VERSION : 0.1
   VAR_INPUT
      IN_xCycleON : Bool;   // Cycle ON
      IN_xCycleONDel : Bool;   // Delayed cycle ON signal
      IN_xResetAlarms : Bool;   // Reset alarms
      IN_xFaultsEnabled : Bool;   // Faults enabled
      IN_xAccelation : Bool;
      IN_rgtMotorConfig : "UDT_MotorConfig";
   END_VAR
   VAR
      ST_xCondOkMan : Bool;   // Manual condition Ok
      ST_xManualMode : Bool;   // Manual mode
      ST_xMachineAnomaly : Bool;   // Machine anomaly
      ST_xStoppingFaults : Bool;   // Stopping fault
      ST_xFaults : Bool;   // Fault
      ST_xWarnings : Bool;   // Warnings
      ST_xConditionOkStopCycle : Bool;   // Condition ok stop cycle
      ST_xOutputEnable : Bool;   // Output enable
      ST_xFeedbackRotation : Bool;   // Feedback rotation
      ST_xPowerUnitSwitchOnRequest : Bool;   // Power unit switch on request
      INPUT_xLocalSwitch : Bool;   // Input local safety switch
      INPUT_xQFMotorFan : Bool;   // Input motor fan protection
      INPUT_xMotorThermalProbe : Bool;   // Input motor thermal probe
      INPUT_xPowerModuleOn : Bool;   // Input power module switched on
      INPUT_dMagnitude : Int;   // Input magnitude value from drive
      INPUT_dTorque : Int;   // Input torque value from drive
      AUX_dReqSpeed_mm_min : DInt := 0;   // Conveyor requested speed [mm/min]
      AUX_dlimitTorqueCorrection : DInt := 0;   // Limit Torque [mm/min]
      tmON_DelayReadyToMove : "UDT_IECTON_V1.00";   // Delay ready to move
      tmON_FeedbackTimeOut : "UDT_IECTON_V1.00";   // Feedback Time out
      tmOF_DriveEnable : "UDT_IECTON_V1.00";   // Drive enable dealy
      AUX_rgtSinamicsIDB : "SINAMICS_LinearPos_ControlTorque";
      tHMR : Struct   // {[Unit]|[Scada Unit]|[LowLimit]|[HigLimit]|[Acces]}
         xManualCommandEnabled : Bool;   // Manual Command enabled {x|x|x|x|O}
         dState : DInt;   // State Conveyor (1=No anomaly, 3=Run, 7=Anomaly) {x|x|x|x|O}
         dMagnitudeCurrent : DInt;   // Magnitude Current [mA] {mA|A|x|x|O}
         dTorque : DInt;   // Torque value [mN] {mN|N|x|x|O}
         dSpeedFeedback : DInt;   // Speed Feedback [mm/min] {mm/min|m/min|x|x|O}
         tManCmd : Struct
            xFdbkRunFw : Bool;   // Motor Rotation Enabled FW {x|x|x|x|O}
         END_STRUCT;
      END_STRUCT;
      tHMW : Struct   // {[Unit]|[Scada Unit]|[LowLimit]|[HigLimit]|[Acces]}
         xEnableManualCommand : Bool;   // Enable Manual command {x|x|x|x|O}
         dSpeedCorrection : DInt;   // Speed Correction[‰] {‰|%|-2|2|M}
         dCurrentLimit : DInt;   // Current limit [‰] {‰|%|0|200|M}
         tManCmd : Struct
            xRunFw : Bool;   // Rotation FW {x|x|x|x|O}
         END_STRUCT;
      END_STRUCT;
      tALM : Struct   // HMI Alarms
         tS : Struct   // Stopping faults
            xLocalSafetySwitch : Bool;   // Local Safety Switch
            xFeedbackError : Bool;   // Feedback Error
            xDriveError : Bool;   // Drive Error
            xMotorFanProtection : Bool;   // Motor Fan protection
            xMotorThermalProbe : Bool;   // Motor Thermal Probe
            xSpare_5 : Bool;
            xSpare_6 : Bool;
            xSpare_7 : Bool;
            xSpare_8 : Bool;
            xSpare_9 : Bool;
            xSpare_10 : Bool;
            xSpare_11 : Bool;
            xSpare_12 : Bool;
            xSpare_13 : Bool;
            xSpare_14 : Bool;
            xSpare_15 : Bool;
            xSpare_16 : Bool;
            xSpare_17 : Bool;
            xSpare_18 : Bool;
            xSpare_19 : Bool;
            xSpare_20 : Bool;
            xSpare_21 : Bool;
            xSpare_22 : Bool;
            xSpare_23 : Bool;
            xSpare_24 : Bool;
            xSpare_25 : Bool;
            xSpare_26 : Bool;
            xSpare_27 : Bool;
            xSpare_28 : Bool;
            xSpare_29 : Bool;
            xSpare_30 : Bool;
            xSpare_31 : Bool;
         END_STRUCT;
         tF : Struct   // Faults
            xSpare_0 : Bool;
            xSpare_1 : Bool;
            xSpare_2 : Bool;
            xSpare_3 : Bool;
            xSpare_4 : Bool;
            xSpare_5 : Bool;
            xSpare_6 : Bool;
            xSpare_7 : Bool;
            xSpare_8 : Bool;
            xSpare_9 : Bool;
            xSpare_10 : Bool;
            xSpare_11 : Bool;
            xSpare_12 : Bool;
            xSpare_13 : Bool;
            xSpare_14 : Bool;
            xSpare_15 : Bool;
            xSpare_16 : Bool;
            xSpare_17 : Bool;
            xSpare_18 : Bool;
            xSpare_19 : Bool;
            xSpare_20 : Bool;
            xSpare_21 : Bool;
            xSpare_22 : Bool;
            xSpare_23 : Bool;
            xSpare_24 : Bool;
            xSpare_25 : Bool;
            xSpare_26 : Bool;
            xSpare_27 : Bool;
            xSpare_28 : Bool;
            xSpare_29 : Bool;
            xSpare_30 : Bool;
            xSpare_31 : Bool;
         END_STRUCT;
         tW : Struct   // Warnings
            xSpare_0 : Bool;
            xSpare_1 : Bool;
            xSpare_2 : Bool;
            xSpare_3 : Bool;
            xSpare_4 : Bool;
            xSpare_5 : Bool;
            xSpare_6 : Bool;
            xSpare_7 : Bool;
            xSpare_8 : Bool;
            xSpare_9 : Bool;
            xSpare_10 : Bool;
            xSpare_11 : Bool;
            xSpare_12 : Bool;
            xSpare_13 : Bool;
            xSpare_14 : Bool;
            xSpare_15 : Bool;
            xSpare_16 : Bool;
            xSpare_17 : Bool;
            xSpare_18 : Bool;
            xSpare_19 : Bool;
            xSpare_20 : Bool;
            xSpare_21 : Bool;
            xSpare_22 : Bool;
            xSpare_23 : Bool;
            xSpare_24 : Bool;
            xSpare_25 : Bool;
            xSpare_26 : Bool;
            xSpare_27 : Bool;
            xSpare_28 : Bool;
            xSpare_29 : Bool;
            xSpare_30 : Bool;
            xSpare_31 : Bool;
         END_STRUCT;
      END_STRUCT;
   END_VAR
   VAR_TEMP
      TMP_dIndex : DInt;
      TMP_dwValue : DWord;
      TMP_iRetVal : Int;
      TMP_xDriveRun : Bool;
      TMP_xDriveEnable : Bool;
   END_VAR
   VAR_TEMP   // added for the SCL form of the ladder/FBD networks
      _w1 : Bool;
   END_VAR
BEGIN

REGION Network 1: #####_MATCH_#####
END_REGION

REGION Network 2: Feedback roller rotation
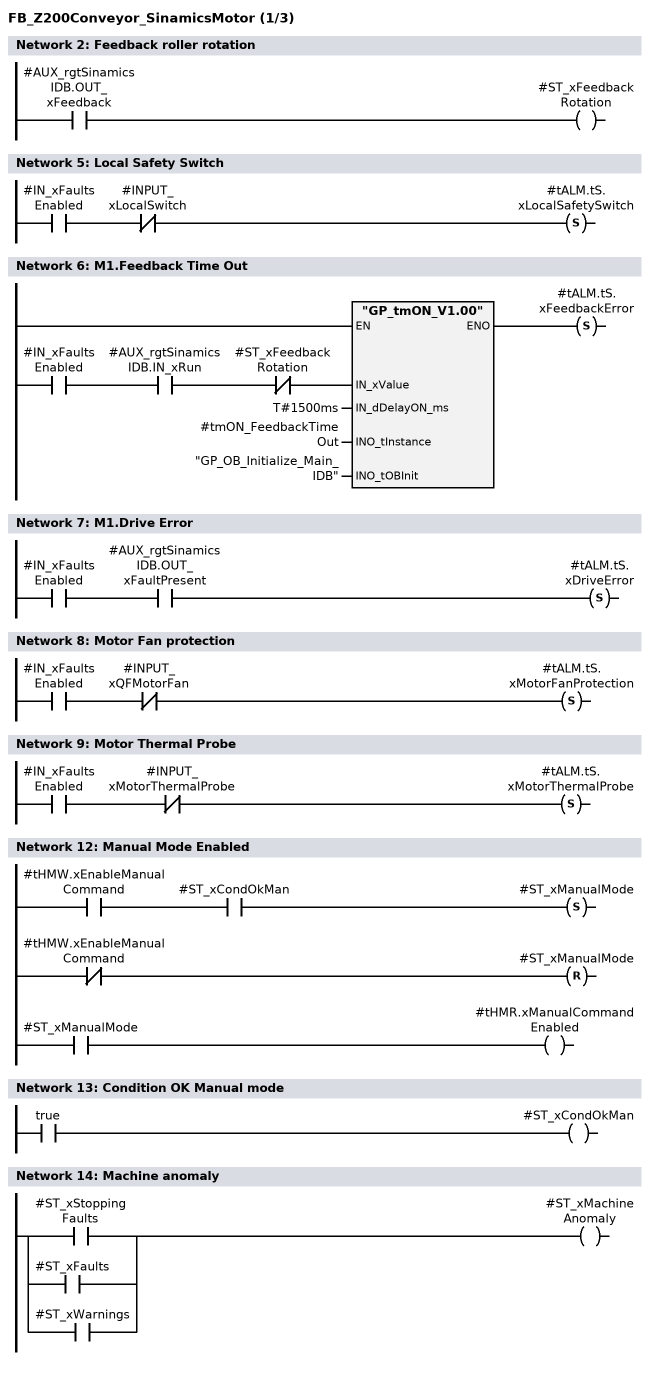
   RUNG wire#powerrail
      Contact( #AUX_rgtSinamicsIDB.OUT_xFeedback )
      Coil( #ST_xFeedbackRotation )
   END_RUNG
   // the same network as SCL:
   #ST_xFeedbackRotation := #AUX_rgtSinamicsIDB.OUT_xFeedback;
END_REGION

REGION Network 3: ####_ALARMS_####
END_REGION

REGION Network 4 (SCL): Reset alarms
   IF #IN_xResetAlarms THEN

       #TMP_dwValue := 0;

       SCATTER(IN:=#TMP_dwValue,
               OUT=>#tALM.tS);

       SCATTER(IN:=#TMP_dwValue,
               OUT=>#tALM.tF);

       SCATTER(IN:=#TMP_dwValue,
               OUT=>#tALM.tW);


   END_IF;
END_REGION

REGION Network 5: Local Safety Switch
   RUNG wire#powerrail
      Contact( #IN_xFaultsEnabled )
      I_Contact( #INPUT_xLocalSwitch )
      S_Coil( #tALM.tS.xLocalSafetySwitch )
   END_RUNG
   // the same network as SCL:
   IF #IN_xFaultsEnabled AND NOT #INPUT_xLocalSwitch THEN #tALM.tS.xLocalSafetySwitch := TRUE; END_IF;
END_REGION

REGION Network 6: M1.Feedback Time Out
   RUNG wire#powerrail
      "GP_tmON_V1.00"(IN_xValue := wire#w1, IN_dDelayON_ms := T#1500ms, INO_tInstance := #tmON_FeedbackTimeOut, INO_tOBInit := "GP_OB_Initialize_Main_IDB")
      S_Coil( #tALM.tS.xFeedbackError )
   END_RUNG
   RUNG wire#powerrail
      Contact( #IN_xFaultsEnabled )
      Contact( #AUX_rgtSinamicsIDB.IN_xRun )
      I_Contact( #ST_xFeedbackRotation )
   END_RUNG wire#w1
   // the same network as SCL:
   "GP_tmON_V1.00"(IN_xValue := #IN_xFaultsEnabled AND #AUX_rgtSinamicsIDB.IN_xRun AND NOT #ST_xFeedbackRotation,
                   IN_dDelayON_ms := T#1500ms,
                   INO_tInstance := #tmON_FeedbackTimeOut,
                   INO_tOBInit := "GP_OB_Initialize_Main_IDB",
                   ENO => #_w1);
   IF #_w1 THEN #tALM.tS.xFeedbackError := TRUE; END_IF;
END_REGION

REGION Network 7: M1.Drive Error
   RUNG wire#powerrail
      Contact( #IN_xFaultsEnabled )
      Contact( #AUX_rgtSinamicsIDB.OUT_xFaultPresent )
      S_Coil( #tALM.tS.xDriveError )
   END_RUNG
   // the same network as SCL:
   IF #IN_xFaultsEnabled AND #AUX_rgtSinamicsIDB.OUT_xFaultPresent THEN #tALM.tS.xDriveError := TRUE; END_IF;
END_REGION

REGION Network 8: Motor Fan protection
   RUNG wire#powerrail
      Contact( #IN_xFaultsEnabled )
      I_Contact( #INPUT_xQFMotorFan )
      S_Coil( #tALM.tS.xMotorFanProtection )
   END_RUNG
   // the same network as SCL:
   IF #IN_xFaultsEnabled AND NOT #INPUT_xQFMotorFan THEN #tALM.tS.xMotorFanProtection := TRUE; END_IF;
END_REGION

REGION Network 9: Motor Thermal Probe
   RUNG wire#powerrail
      Contact( #IN_xFaultsEnabled )
      I_Contact( #INPUT_xMotorThermalProbe )
      S_Coil( #tALM.tS.xMotorThermalProbe )
   END_RUNG
   // the same network as SCL:
   IF #IN_xFaultsEnabled AND NOT #INPUT_xMotorThermalProbe THEN #tALM.tS.xMotorThermalProbe := TRUE; END_IF;
END_REGION

REGION Network 10 (SCL): Calculate general statuses
   GATHER(IN:=#tALM.tS,
          OUT=>#TMP_dwValue);

   IF #TMP_dwValue <> 0 THEN
       #ST_xStoppingFaults := TRUE;
   ELSE
       #ST_xStoppingFaults := FALSE;
   END_IF;

   GATHER(IN:=#tALM.tF,
          OUT=>#TMP_dwValue);

   IF #TMP_dwValue <> 0 THEN
       #ST_xFaults := TRUE;
   ELSE
       #ST_xFaults := FALSE;
   END_IF;

   GATHER(IN:=#tALM.tW,
          OUT=>#TMP_dwValue);

   IF #TMP_dwValue <> 0 THEN
       #ST_xWarnings := TRUE;
   ELSE
       #ST_xWarnings := FALSE;
   END_IF;
END_REGION

REGION Network 11: #####_HMI_LOGICS_#####
END_REGION

REGION Network 12: Manual Mode Enabled
   RUNG wire#powerrail
      Contact( #tHMW.xEnableManualCommand )
      Contact( #ST_xCondOkMan )
      S_Coil( #ST_xManualMode )
   END_RUNG
   RUNG wire#powerrail
      I_Contact( #tHMW.xEnableManualCommand )
      R_Coil( #ST_xManualMode )
   END_RUNG
   RUNG wire#powerrail
      Contact( #ST_xManualMode )
      Coil( #tHMR.xManualCommandEnabled )
   END_RUNG
   // the same network as SCL:
   IF #tHMW.xEnableManualCommand AND #ST_xCondOkMan THEN #ST_xManualMode := TRUE; END_IF;
   IF NOT #tHMW.xEnableManualCommand THEN #ST_xManualMode := FALSE; END_IF;
   #tHMR.xManualCommandEnabled := #ST_xManualMode;
END_REGION

REGION Network 13: Condition OK Manual mode
   RUNG wire#powerrail
      Contact( true )
      Coil( #ST_xCondOkMan )
   END_RUNG
   // the same network as SCL:
   #ST_xCondOkMan := true;
END_REGION

REGION Network 14: Machine anomaly
   RUNG wire#powerrail
      Contact( #ST_xStoppingFaults )
      wire#w1
      Coil( #ST_xMachineAnomaly )
   END_RUNG
   RUNG wire#powerrail
      Contact( #ST_xFaults )
   END_RUNG wire#w1
   RUNG wire#powerrail
      Contact( #ST_xWarnings )
   END_RUNG wire#w1
   // the same network as SCL:
   #ST_xMachineAnomaly := #ST_xStoppingFaults OR #ST_xFaults OR #ST_xWarnings;
END_REGION

REGION Network 15: Output Enable
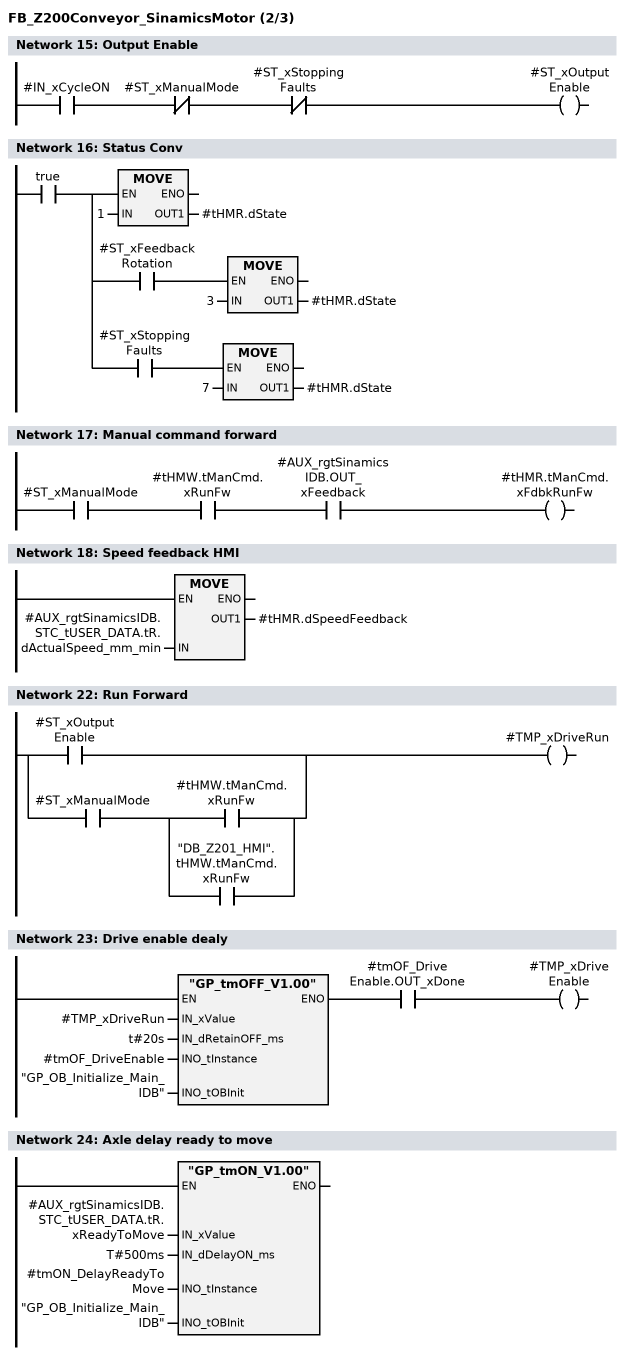
   RUNG wire#powerrail
      Contact( #IN_xCycleON )
      I_Contact( #ST_xManualMode )
      I_Contact( #ST_xStoppingFaults )
      Coil( #ST_xOutputEnable )
   END_RUNG
   // the same network as SCL:
   #ST_xOutputEnable := #IN_xCycleON AND NOT #ST_xManualMode AND NOT #ST_xStoppingFaults;
END_REGION

REGION Network 16: Status Conv
   RUNG wire#powerrail
      Contact( true )
      wire#w1
      Move(in := 1, out1 => #tHMR.dState)
   END_RUNG
   RUNG wire#w1
      Contact( #ST_xFeedbackRotation )
      Move(in := 3, out1 => #tHMR.dState)
   END_RUNG
   RUNG wire#w1
      Contact( #ST_xStoppingFaults )
      Move(in := 7, out1 => #tHMR.dState)
   END_RUNG
   // the same network as SCL:
   IF true THEN #tHMR.dState := 1; END_IF;
   IF true AND #ST_xFeedbackRotation THEN #tHMR.dState := 3; END_IF;
   IF true AND #ST_xStoppingFaults THEN #tHMR.dState := 7; END_IF;
END_REGION

REGION Network 17: Manual command forward
   RUNG wire#powerrail
      Contact( #ST_xManualMode )
      Contact( #tHMW.tManCmd.xRunFw )
      Contact( #AUX_rgtSinamicsIDB.OUT_xFeedback )
      Coil( #tHMR.tManCmd.xFdbkRunFw )
   END_RUNG
   // the same network as SCL:
   #tHMR.tManCmd.xFdbkRunFw := #ST_xManualMode AND #tHMW.tManCmd.xRunFw AND #AUX_rgtSinamicsIDB.OUT_xFeedback;
END_REGION

REGION Network 18: Speed feedback HMI
   RUNG wire#powerrail
      Move(in := #AUX_rgtSinamicsIDB.STC_tUSER_DATA.tR.dActualSpeed_mm_min, out1 => #tHMR.dSpeedFeedback)
   END_RUNG
   // the same network as SCL:
   #tHMR.dSpeedFeedback := #AUX_rgtSinamicsIDB.STC_tUSER_DATA.tR.dActualSpeed_mm_min;
END_REGION

REGION Network 19 (SCL): Torque and current feedback
   #tHMR.dMagnitudeCurrent := LREAL_TO_DINT(9.6 / 16384.0 * #INPUT_dMagnitude * 1000);
   #tHMR.dTorque := LREAL_TO_DINT(28.8 / 16384.0 * #INPUT_dTorque * 1000);
END_REGION

REGION Network 20: #####_OUTPUT_#####
END_REGION

REGION Network 21 (SCL): Constant
   //####,#Motor Costant#####
   //Adrress of Synamisc Motor
   #AUX_rgtSinamicsIDB.STC_tSYS_DATA.iIOAddress_MM := #IN_rgtMotorConfig.iIOAddress_MM;
   //Type of telegram(1=Open/closeLoop;111=Positioning)
   #AUX_rgtSinamicsIDB.STC_tSYS_DATA.iPZD_MM := #IN_rgtMotorConfig.iPZD_MM;
   //Max Speed (set equal to StarterProject)[Rpm]
   #AUX_rgtSinamicsIDB.STC_tSYS_DATA.dMaxSpeed_rpm := #IN_rgtMotorConfig.dMaxSpeed_rpm;
   //K Conversion From RPM to mm/min (value come from Drive)
   #AUX_rgtSinamicsIDB.STC_tSYS_DATA.rK_rpm_mmMin := #IN_rgtMotorConfig.rK_rpm_mmMin;
   //K Conversion From mm/min to Rpm (for Open Close Loop) value for Drive
   #AUX_rgtSinamicsIDB.STC_tSYS_DATA.rK_mmMin_Rpm := #IN_rgtMotorConfig.rK_mmMin_Rpm;
   //Max Acceleration [Pos=m/s2, OpnLoop=S]
   #AUX_rgtSinamicsIDB.STC_tSYS_DATA.rMaxAcc := #IN_rgtMotorConfig.rMaxAcc;
   //Max Deceleration [Pos=m/s2, OpnLoop=S]
   #AUX_rgtSinamicsIDB.STC_tSYS_DATA.rMaxDec := #IN_rgtMotorConfig.rMaxDec;
   //Ramp Value Acceleration [Pos=m/s2, OpnLoop=S]
   #AUX_rgtSinamicsIDB.STC_tUSER_DATA.tW.rAcc := #IN_rgtMotorConfig.rAcc;
   //Ramp Value Deceleration [Pos=m/s2, OpnLoop=S]
   #AUX_rgtSinamicsIDB.STC_tUSER_DATA.tW.rDec := #IN_rgtMotorConfig.rDec;
   //Enable Module Correction
   #AUX_rgtSinamicsIDB.STC_tEXT_DATA.tW.xModuleCorrect := #IN_rgtMotorConfig.xModuleCorrect;
   //MDI
   #AUX_rgtSinamicsIDB.STC_tUSER_DATA.tW.xMDI_Continue := #IN_rgtMotorConfig.xMDI_Continue;
END_REGION

REGION Network 22: Run Forward
   RUNG wire#powerrail
      Contact( #ST_xOutputEnable )
      wire#w1
      Coil( #TMP_xDriveRun )
   END_RUNG
   RUNG wire#powerrail
      Contact( #ST_xManualMode )
      wire#w2
      Contact( #tHMW.tManCmd.xRunFw )
   END_RUNG wire#w1
   RUNG wire#w2
      Contact( "DB_Z201_HMI".tHMW.tManCmd.xRunFw )
   END_RUNG wire#w1
   // the same network as SCL:
   #TMP_xDriveRun := #ST_xOutputEnable OR (#ST_xManualMode AND (#tHMW.tManCmd.xRunFw OR "DB_Z201_HMI".tHMW.tManCmd.xRunFw));
END_REGION

REGION Network 23: Drive enable dealy
   RUNG wire#powerrail
      "GP_tmOFF_V1.00"(IN_xValue := #TMP_xDriveRun, IN_dRetainOFF_ms := t#20s, INO_tInstance := #tmOF_DriveEnable, INO_tOBInit := "GP_OB_Initialize_Main_IDB")
      Contact( #tmOF_DriveEnable.OUT_xDone )
      Coil( #TMP_xDriveEnable )
   END_RUNG
   // the same network as SCL:
   "GP_tmOFF_V1.00"(IN_xValue := #TMP_xDriveRun,
                    IN_dRetainOFF_ms := t#20s,
                    INO_tInstance := #tmOF_DriveEnable,
                    INO_tOBInit := "GP_OB_Initialize_Main_IDB",
                    ENO => #_w1);
   #TMP_xDriveEnable := #_w1 AND #tmOF_DriveEnable.OUT_xDone;
END_REGION

REGION Network 24: Axle delay ready to move
   RUNG wire#powerrail
      "GP_tmON_V1.00"(IN_xValue := #AUX_rgtSinamicsIDB.STC_tUSER_DATA.tR.xReadyToMove, IN_dDelayON_ms := T#500ms, INO_tInstance := #tmON_DelayReadyToMove, INO_tOBInit := "GP_OB_Initialize_Main_IDB")
   END_RUNG
   // the same network as SCL:
   "GP_tmON_V1.00"(IN_xValue := #AUX_rgtSinamicsIDB.STC_tUSER_DATA.tR.xReadyToMove,
                   IN_dDelayON_ms := T#500ms,
                   INO_tInstance := #tmON_DelayReadyToMove,
                   INO_tOBInit := "GP_OB_Initialize_Main_IDB");
END_REGION

REGION Network 25: Timer done
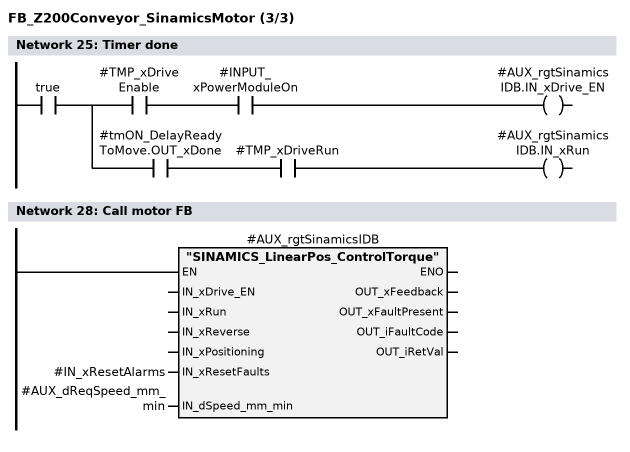
   RUNG wire#powerrail
      Contact( true )
      wire#w1
      Contact( #TMP_xDriveEnable )
      Contact( #INPUT_xPowerModuleOn )
      Coil( #AUX_rgtSinamicsIDB.IN_xDrive_EN )
   END_RUNG
   RUNG wire#w1
      Contact( #tmON_DelayReadyToMove.OUT_xDone )
      Contact( #TMP_xDriveRun )
      Coil( #AUX_rgtSinamicsIDB.IN_xRun )
   END_RUNG
   // the same network as SCL:
   #AUX_rgtSinamicsIDB.IN_xDrive_EN := true AND #TMP_xDriveEnable AND #INPUT_xPowerModuleOn;
   #AUX_rgtSinamicsIDB.IN_xRun := true AND #tmON_DelayReadyToMove.OUT_xDone AND #TMP_xDriveRun;
END_REGION

REGION Network 26 (SCL): Manager Speed
   IF #IN_xAccelation = FALSE THEN
       #AUX_dReqSpeed_mm_min :="FB_LehrSpeed_IDB".tHMR.dActualSpeedValueToConveyor_mm_min * ((#tHMW.dSpeedCorrection + 1000) / 1000);
   ELSE
       #AUX_dReqSpeed_mm_min := "FB_LehrSpeed_IDB".tHMR.dActualSpeedValueToConveyor_mm_min + 20000;
   END_IF;
END_REGION

REGION Network 27 (SCL): Limit Torque
   #AUX_dlimitTorqueCorrection := REAL_TO_DINT((DINT_TO_REAL(#tHMW.dCurrentLimit) / 2000.0) * 16384.0);
   #AUX_rgtSinamicsIDB.STC_tPZD_OpCLLoop.tW.iTorque := DINT_TO_INT(#AUX_dlimitTorqueCorrection);
END_REGION

REGION Network 28: Call motor FB
   RUNG wire#powerrail
      #AUX_rgtSinamicsIDB(IN_xDrive_EN :=, IN_xRun :=, IN_xReverse :=, IN_xPositioning :=, IN_xResetFaults := #IN_xResetAlarms, IN_dSpeed_mm_min := #AUX_dReqSpeed_mm_min, OUT_xFeedback =>, OUT_xFaultPresent =>, OUT_iFaultCode =>, OUT_iRetVal =>)
   END_RUNG
   // the same network as SCL:
   #AUX_rgtSinamicsIDB(IN_xResetFaults := #IN_xResetAlarms, IN_dSpeed_mm_min := #AUX_dReqSpeed_mm_min);   // "SINAMICS_LinearPos_ControlTorque"
END_REGION
END_FUNCTION_BLOCK

FUNCTION "Z200SinamicsCU_Management" : Void   // FC115, LAD
{ S7_Optimized_Access := 'TRUE' }
VERSION : 0.1
BEGIN

REGION Network 1: ###############_A250AP1_##############
END_REGION

REGION Network 2 (SCL): Mapping
   "CU_A250AP1_IDB".STC_tSYS_DATA.iIOAddress_CU := 2000;
   "CU_A250AP1_IDB".STC_tSYS_DATA.iIOAddress_PM :=2010;
   "CU_A250AP1_IDB".STC_tSYS_DATA.iPowerOFFDelay_ms := 3000;
END_REGION

REGION Network 3: CU
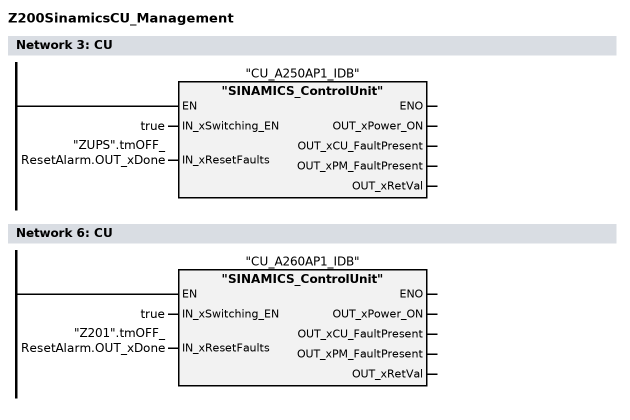
   RUNG wire#powerrail
      "CU_A250AP1_IDB"(IN_xSwitching_EN := true, IN_xResetFaults := "ZUPS".tmOFF_ResetAlarm.OUT_xDone, OUT_xPower_ON =>, OUT_xCU_FaultPresent =>, OUT_xPM_FaultPresent =>, OUT_xRetVal =>)
   END_RUNG
   // the same network as SCL:
   "CU_A250AP1_IDB"(IN_xSwitching_EN := true, IN_xResetFaults := "ZUPS".tmOFF_ResetAlarm.OUT_xDone);   // "SINAMICS_ControlUnit"
END_REGION

REGION Network 4: ###############_A260AP1_############## / ###############_A102AP1_##############
END_REGION

REGION Network 5 (SCL): Mapping
   "CU_A260AP1_IDB".STC_tSYS_DATA.iIOAddress_CU := 2200;
   "CU_A260AP1_IDB".STC_tSYS_DATA.iIOAddress_PM :=2210;
   "CU_A260AP1_IDB".STC_tSYS_DATA.iPowerOFFDelay_ms := 3000;
END_REGION

REGION Network 6: CU
   RUNG wire#powerrail
      "CU_A260AP1_IDB"(IN_xSwitching_EN := true, IN_xResetFaults := "Z201".tmOFF_ResetAlarm.OUT_xDone, OUT_xPower_ON =>, OUT_xCU_FaultPresent =>, OUT_xPM_FaultPresent =>, OUT_xRetVal =>)
   END_RUNG
   // the same network as SCL:
   "CU_A260AP1_IDB"(IN_xSwitching_EN := true, IN_xResetFaults := "Z201".tmOFF_ResetAlarm.OUT_xDone);   // "SINAMICS_ControlUnit"
END_REGION
END_FUNCTION

// folder: 03_Programs_Logics/MCC1201/27_T1DropConveyor

FUNCTION_BLOCK "FB_DropConveyor"   // FB23, LAD
{ S7_Optimized_Access := 'TRUE' }
VERSION : 0.1
   VAR_INPUT
      IN_xCycleON : Bool;   // Cycle ON
      IN_xCycleONDel : Bool;   // Delayed cycle ON signal
      IN_xManualMode : Bool;   // Manual mode drop conveyor
      IN_xResetAlarms : Bool;   // Reset alarms
      IN_xFaultsEnabled : Bool;   // Faults enabled
      IN_dGlassBreakMachineIndex : DInt;   // Glass break machine index
      IN_dGlassBreakGetIndex : DInt;   // Glass break get index
      IN_dActualLehrSpeed_mm_min : DInt;   // Lehr speed (mm/min)
      IN_xSimulationActive : Bool;   // Enable simulation (EXPERT USER)
      INPUT : Struct
         xProtection : Bool := false;   // Input.Protection motor
         xProtectionBrake : Bool := false;   // Input.Protection brake
         xFeedbackMovement : Bool := false;   // Input.Movement feedback
         xSafetyBar : Bool := false;   // Input.Safety bar inserted
         xDoorOpen : Bool := false;   // Input.Door open
         xUpPosition : Bool := false;   // Input.Up position
         xDownPosition : Bool := false;   // Input.Down position
         xUpDownPushbutton : Bool := false;   // Input.Up/Down pushbutton
      END_STRUCT;
   END_VAR
   VAR_OUTPUT
      OUTPUT : Struct
         xRiseDrop : Bool := false;   // Output.Rise drop conveyor
         xDescentDrop : Bool := false;   // Output.Descent drop conveyor
         xHLDoorOpen : Bool;
         xHLUpDownPushbutton : Bool := false;   // Output.HL Up/Down pushbutton
      END_STRUCT;
   END_VAR
   VAR_IN_OUT
      INO_tRibbon : "UDT_RibbonData";   // Ribbon data
   END_VAR
   VAR
      ST_xPhaseInProgress : Bool := false;   // Phase in progress
      ST_xFaults : Bool := false;   // Cumulative of faults
      ST_xStoppingFaults : Bool := false;   // Cumulative of stopping faults
      ST_xWarnings : Bool := false;   // Cumulative of warning
      AUX_tmONFeedbackAlarm : TON_TIME;   // Feedback alarm
      AUX_tmONMismatchSensorAlarm : TON_TIME;   // Mismatch sensor feedback alarm
      AUX_tmONUpSensorAlarm : TON_TIME;   // Up sensor feedback alarm
      AUX_tmONDownSensorAlarm : TON_TIME;   // Down sensor feedback alarm
      AUX_tmONForceUp : TON_TIME;   // Force up
      ST_xConditionOKforStopCycle : Bool := false;   // Condition for stop cycle
      ST_xConveyorUpRequest : Bool := false;   // Conveyor Up request
      ST_xConveyorDwRequest : Bool := false;   // Conveyor Down request
      ST_xConveyorUp : Bool := false;   // Conveyor Up
      ST_xUpFromPush : Bool := false;   // Up from pushbutton
      ST_xOutputEnable : Bool := false;   // Output enable
      ST_xUpFromScada : Bool := false;   // Up from scada
      ST_xGlassBreak : Bool;   // Glass break under bridge
      OSR_xChangeState : Bool;   // OSR change state report
      OSR_xConditionOk : Bool;   // OSR condition ok report
      OSR_xConditionNotOk : Bool;   // OSR condition not ok report
      OSR_xMemoryState : Bool;   // OSR memory state report
      OSN_xMemory : Bool;   // OSN memory report
      OSR_xUpDownSBRequest : Bool := false;   // OSR Up/Down pushbutton request
      OS_xUpDownSBRequest : Bool := false;   // OS Up/Down pushbutton request
      OSR_xForceUpSBRequest : Bool := false;   // OSR force up pushbutton request
      OS_xForceUpSBRequest : Bool := false;   // OS force up pushbutton request
      OSR_xRise : Bool := false;   // OSR Rise
      OS_xRise : Bool := false;   // OS Rise
      OSR_xDescent : Bool := false;   // OSR Descent
      OS_xDescent : Bool := false;   // OS Descent
      OSR_xManCmdRise : Bool := false;   // OSR Man Cmd Rise
      OS_xManCmdRise : Bool := false;   // OS Man Cmd Rise
      OSR_xManCmdDescent : Bool := false;   // OSR Man Cmd Descent
      OS_xManCmdDescent : Bool := false;   // OS Man Cmd Descent
      OSR_xBreak : Bool := false;   // OSR Glass break
   END_VAR
   VAR RETAIN
      tHMW : Struct   // HMI Write
         tManCmd : Struct
            xRise : Bool := false;   // Manual rise {x|x|x|x|O}
            xDescent : Bool := false;   // Manual descent {x|x|x|x|O}
         END_STRUCT;
         dDistanceFromSnaproll_cmm : DInt;   // Distance from snaproll [mm/100] {mm/100|mm|0|65000|M}
         xUpdateDistanceFromSnaproll : Bool;   // Update distance from snaproll {x|x|x|x|M}
         xEnabledBreakingDetection : Bool;   // Enable automatic descent for glass break {x|x|x|x|O}
         xRequestUp : Bool;   // Request tilting up {x|x|x|x|M}
         xRequestDown : Bool;   // Request tilting down {x|x|x|x|M}
         xForceUp : Bool;   // Force tilting up {x|x|x|x|M}
         xForceDown : Bool;   // Force tilting down {x|x|x|x|M}
      END_STRUCT;
      tHMR : Struct   // HMI Read
         tManCmd : Struct
            xRiseFdbk : Bool;   // Manual rise fdbk {x|x|x|x|O}
            xDescentFdbk : Bool;   // Manual descent fdbk {x|x|x|x|O}
         END_STRUCT;
         xUpPosition : Bool;   // Up position {x|x|x|x|O}
         xDownPosition : Bool;   // Down position {x|x|x|x|O}
         dMode : DInt;   // Drop mode (1=Down 2=Up 4=Req Down 8=Req up)
         dStatus : DInt;   // Conveyor status (1=Idle 3=Running 7=Anomaly)
         dDistanceFromSnaproll_cmm : DInt;   // Distance from snaproll [mm/100] {mm/100|mm|x|x|O}
      END_STRUCT;
   END_VAR
   VAR
      tALM : Struct   // HMI Alarms
         tW : Struct   // Warnings
            xDoorOpen : Bool;   // Door open
            xSpare_1 : Bool;
            xSpare_2 : Bool;
            xSpare_3 : Bool;
            xSpare_4 : Bool;
            xSpare_5 : Bool;
            xSpare_6 : Bool;
            xSpare_7 : Bool;
            xSpare_8 : Bool;
            xSpare_9 : Bool;
            xSpare_10 : Bool;
            xSpare_11 : Bool;
            xSpare_12 : Bool;
            xSpare_13 : Bool;
            xSpare_14 : Bool;
            xSpare_15 : Bool;
            xSpare_16 : Bool;
            xSpare_17 : Bool;
            xSpare_18 : Bool;
            xSpare_19 : Bool;
            xSpare_20 : Bool;
            xSpare_21 : Bool;
            xSpare_22 : Bool;
            xSpare_23 : Bool;
            xSpare_24 : Bool;
            xSpare_25 : Bool;
            xSpare_26 : Bool;
            xSpare_27 : Bool;
            xSpare_28 : Bool;
            xSpare_29 : Bool;
            xSpare_30 : Bool;
            xSpare_31 : Bool;
         END_STRUCT;
         tF : Struct   // Faults
            xSpare_0 : Bool;
            xSpare_1 : Bool;
            xSpare_2 : Bool;
            xSpare_3 : Bool;
            xSpare_4 : Bool;
            xSpare_5 : Bool;
            xSpare_6 : Bool;
            xSpare_7 : Bool;
            xSpare_8 : Bool;
            xSpare_9 : Bool;
            xSpare_10 : Bool;
            xSpare_11 : Bool;
            xSpare_12 : Bool;
            xSpare_13 : Bool;
            xSpare_14 : Bool;
            xSpare_15 : Bool;
            xSpare_16 : Bool;
            xSpare_17 : Bool;
            xSpare_18 : Bool;
            xSpare_19 : Bool;
            xSpare_20 : Bool;
            xSpare_21 : Bool;
            xSpare_22 : Bool;
            xSpare_23 : Bool;
            xSpare_24 : Bool;
            xSpare_25 : Bool;
            xSpare_26 : Bool;
            xSpare_27 : Bool;
            xSpare_28 : Bool;
            xSpare_29 : Bool;
            xSpare_30 : Bool;
            xSpare_31 : Bool;
         END_STRUCT;
         tS : Struct   // Stopping faults
            xProtectionLifting : Bool;   // QM.Protection lifting
            xFeedbackLifting : Bool;   // KM.Feedback lifting
            xTimeoutFrameHigh : Bool;   // SQ.Timeout frame high
            xTimeoutFrameLow : Bool;   // SQ.Timeout frame low
            xSensorsMismatch : Bool;   // SQ.Sensors High/low same status
            xProtectionBrake : Bool;   // QM.Protection brake
            xTiltingSafety : Bool;   // SQ.Safety bar inserted
            xSpare_7 : Bool;
            xSpare_8 : Bool;
            xSpare_9 : Bool;
            xSpare_10 : Bool;
            xSpare_11 : Bool;
            xSpare_12 : Bool;
            xSpare_13 : Bool;
            xSpare_14 : Bool;
            xSpare_15 : Bool;
            xSpare_16 : Bool;
            xSpare_17 : Bool;
            xSpare_18 : Bool;
            xSpare_19 : Bool;
            xSpare_20 : Bool;
            xSpare_21 : Bool;
            xSpare_22 : Bool;
            xSpare_23 : Bool;
            xSpare_24 : Bool;
            xSpare_25 : Bool;
            xSpare_26 : Bool;
            xSpare_27 : Bool;
            xSpare_28 : Bool;
            xSpare_29 : Bool;
            xSpare_30 : Bool;
            xSpare_31 : Bool;
         END_STRUCT;
      END_STRUCT;
   END_VAR
   VAR_TEMP
      TMP_dwValue : DWord;
      TMP_xDummy : Bool;
      TMP_xUpdate : Bool;
      TMP_xError : Bool;
   END_VAR
   VAR CONSTANT
      CONST_DBREAKUPOFF_CMM : DInt := 10000;   // Break upstream offset [mm/100]
      CONST_DBREAKDOWNOFF_CMM : DInt := 10000;   // Break downstream offset [mm/100]
      dDESTINATION_ID_T1 : DInt := 200;
      dSTATUSIDEN_TrapUp : DInt := 21;
      dSTATUSIDEN_TrapDw : DInt := 20;
   END_VAR
   VAR_TEMP   // added for the SCL form of the ladder/FBD networks
      _w1 : Bool;
      _w2 : Bool;
   END_VAR
BEGIN

REGION Network 1 (SCL): ### COSTANTS ###
END_REGION

REGION Network 2: ### MATCH ###
END_REGION

REGION Network 3 (SCL)
   IF #IN_xSimulationActive THEN
       #INPUT.xProtection := 1;
       #INPUT.xProtectionBrake := 1;
       #INPUT.xFeedbackMovement := #OUTPUT.xDescentDrop OR #OUTPUT.xRiseDrop;
       #INPUT.xSafetyBar := 1;
       #INPUT.xDoorOpen := 1;
       IF #tHMR.dMode = 1 OR #tHMR.dMode = 4 THEN
           #INPUT.xUpPosition := 0;
           #INPUT.xDownPosition := 1;
       END_IF;
       IF #tHMR.dMode = 2 OR #tHMR.dMode = 8 THEN
           #INPUT.xDownPosition := 0;
           #INPUT.xUpPosition := 1;
       END_IF;
       IF  NOT #INPUT.xDownPosition AND NOT #INPUT.xUpPosition THEN
           #INPUT.xDownPosition := 1;
           #INPUT.xUpPosition := 0;
       END_IF;
   END_IF;
END_REGION

REGION Network 4: Up down SB request
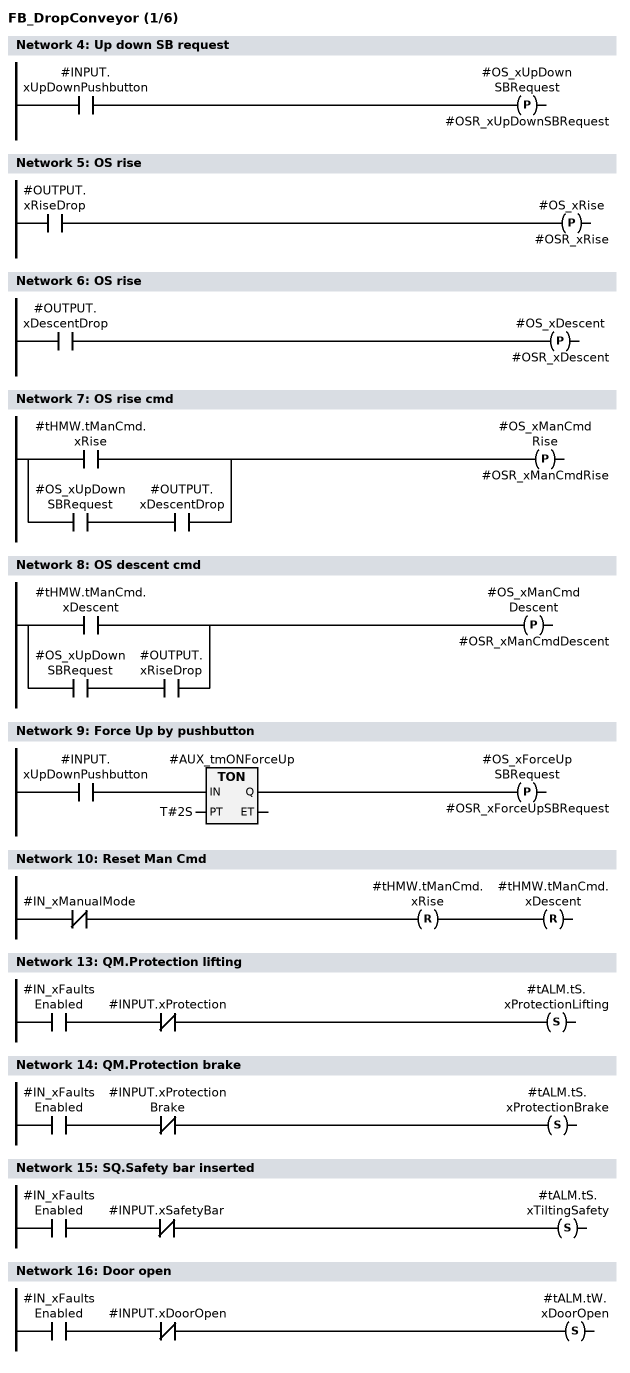
   #OS_xUpDownSBRequest := #INPUT.xUpDownPushbutton AND NOT #OSR_xUpDownSBRequest;   // rising edge
   #OSR_xUpDownSBRequest := #INPUT.xUpDownPushbutton;
END_REGION

REGION Network 5: OS rise
   #OS_xRise := #OUTPUT.xRiseDrop AND NOT #OSR_xRise;   // rising edge
   #OSR_xRise := #OUTPUT.xRiseDrop;
END_REGION

REGION Network 6: OS rise
   #OS_xDescent := #OUTPUT.xDescentDrop AND NOT #OSR_xDescent;   // rising edge
   #OSR_xDescent := #OUTPUT.xDescentDrop;
END_REGION

REGION Network 7: OS rise cmd
   #_w1 := #tHMW.tManCmd.xRise OR (#OS_xUpDownSBRequest AND #OUTPUT.xDescentDrop);
   #OS_xManCmdRise := #_w1 AND NOT #OSR_xManCmdRise;   // rising edge
   #OSR_xManCmdRise := #_w1;
END_REGION

REGION Network 8: OS descent cmd
   #_w1 := #tHMW.tManCmd.xDescent OR (#OS_xUpDownSBRequest AND #OUTPUT.xRiseDrop);
   #OS_xManCmdDescent := #_w1 AND NOT #OSR_xManCmdDescent;   // rising edge
   #OSR_xManCmdDescent := #_w1;
END_REGION

REGION Network 9: Force Up by pushbutton
   #AUX_tmONForceUp(IN := #INPUT.xUpDownPushbutton, PT := T#2S);   // TON
   #OS_xForceUpSBRequest := #AUX_tmONForceUp.Q AND NOT #OSR_xForceUpSBRequest;   // rising edge
   #OSR_xForceUpSBRequest := #AUX_tmONForceUp.Q;
END_REGION

REGION Network 10: Reset Man Cmd
   RUNG wire#powerrail
      I_Contact( #IN_xManualMode )
      R_Coil( #tHMW.tManCmd.xRise )
      R_Coil( #tHMW.tManCmd.xDescent )
   END_RUNG
   // the same network as SCL:
   IF NOT #IN_xManualMode THEN
       #tHMW.tManCmd.xRise := FALSE;
       #tHMW.tManCmd.xDescent := FALSE;
   END_IF;
END_REGION

REGION Network 11: ####_ALARMS_####
END_REGION

REGION Network 12 (SCL): Reset alarms
   IF #IN_xResetAlarms THEN

       #TMP_dwValue := 0;

       SCATTER(IN:=#TMP_dwValue,
               OUT=>#tALM.tS);

       SCATTER(IN:=#TMP_dwValue,
               OUT=>#tALM.tF);

       SCATTER(IN:=#TMP_dwValue,
               OUT=>#tALM.tW);

   END_IF;
END_REGION

REGION Network 13: QM.Protection lifting
   RUNG wire#powerrail
      Contact( #IN_xFaultsEnabled )
      I_Contact( #INPUT.xProtection )
      S_Coil( #tALM.tS.xProtectionLifting )
   END_RUNG
   // the same network as SCL:
   IF #IN_xFaultsEnabled AND NOT #INPUT.xProtection THEN #tALM.tS.xProtectionLifting := TRUE; END_IF;
END_REGION

REGION Network 14: QM.Protection brake
   RUNG wire#powerrail
      Contact( #IN_xFaultsEnabled )
      I_Contact( #INPUT.xProtectionBrake )
      S_Coil( #tALM.tS.xProtectionBrake )
   END_RUNG
   // the same network as SCL:
   IF #IN_xFaultsEnabled AND NOT #INPUT.xProtectionBrake THEN #tALM.tS.xProtectionBrake := TRUE; END_IF;
END_REGION

REGION Network 15: SQ.Safety bar inserted
   RUNG wire#powerrail
      Contact( #IN_xFaultsEnabled )
      I_Contact( #INPUT.xSafetyBar )
      S_Coil( #tALM.tS.xTiltingSafety )
   END_RUNG
   // the same network as SCL:
   IF #IN_xFaultsEnabled AND NOT #INPUT.xSafetyBar THEN #tALM.tS.xTiltingSafety := TRUE; END_IF;
END_REGION

REGION Network 16: Door open
   RUNG wire#powerrail
      Contact( #IN_xFaultsEnabled )
      I_Contact( #INPUT.xDoorOpen )
      S_Coil( #tALM.tW.xDoorOpen )
   END_RUNG
   // the same network as SCL:
   IF #IN_xFaultsEnabled AND NOT #INPUT.xDoorOpen THEN #tALM.tW.xDoorOpen := TRUE; END_IF;
END_REGION

REGION Network 17: KM.Feedback lifting